// TIA Portal project "EMS" (V15.1) (continued)
   "SDC_EMS01_CARRIER61_Spare2" AT %Q6828.2 : Bool;
   "SDC_EMS01_CARRIER61_PositioningComplete" AT %Q6828.3 : Bool;
   "SDC_EMS01_CARRIER61_RunStopPressed" AT %Q6828.4 : Bool;
   "SDC_EMS01_CARRIER61_Moving" AT %Q6828.5 : Bool;
   "SDC_EMS01_CARRIER61_Faulted" AT %Q6828.6 : Bool;
   "SDC_EMS01_CARRIER61_InAuto" AT %Q6828.7 : Bool;
   "SDC_EMS01_CARRIER62_Spare0" AT %Q6829.0 : Bool;
   "SDC_EMS01_CARRIER62_DriveTripped" AT %Q6829.1 : Bool;
   "SDC_EMS01_CARRIER62_Spare2" AT %Q6829.2 : Bool;
   "SDC_EMS01_CARRIER62_PositioningComplete" AT %Q6829.3 : Bool;
   "SDC_EMS01_CARRIER62_RunStopPressed" AT %Q6829.4 : Bool;
   "SDC_EMS01_CARRIER62_Moving" AT %Q6829.5 : Bool;
   "SDC_EMS01_CARRIER62_Faulted" AT %Q6829.6 : Bool;
   "SDC_EMS01_CARRIER62_InAuto" AT %Q6829.7 : Bool;
   "SDC_EMS01_CARRIER63_Spare0" AT %Q6830.0 : Bool;
   "SDC_EMS01_CARRIER63_DriveTripped" AT %Q6830.1 : Bool;
   "SDC_EMS01_CARRIER63_Spare2" AT %Q6830.2 : Bool;
   "SDC_EMS01_CARRIER63_PositioningComplete" AT %Q6830.3 : Bool;
   "SDC_EMS01_CARRIER63_RunStopPressed" AT %Q6830.4 : Bool;
   "SDC_EMS01_CARRIER63_Moving" AT %Q6830.5 : Bool;
   "SDC_EMS01_CARRIER63_Faulted" AT %Q6830.6 : Bool;
   "SDC_EMS01_CARRIER63_InAuto" AT %Q6830.7 : Bool;
   "SDC_EMS01_CARRIER64_Spare0" AT %Q6831.0 : Bool;
   "SDC_EMS01_CARRIER64_DriveTripped" AT %Q6831.1 : Bool;
   "SDC_EMS01_CARRIER64_Spare2" AT %Q6831.2 : Bool;
   "SDC_EMS01_CARRIER64_PositioningComplete" AT %Q6831.3 : Bool;
   "SDC_EMS01_CARRIER64_RunStopPressed" AT %Q6831.4 : Bool;
   "SDC_EMS01_CARRIER64_Moving" AT %Q6831.5 : Bool;
   "SDC_EMS01_CARRIER64_Faulted" AT %Q6831.6 : Bool;
   "SDC_EMS01_CARRIER64_InAuto" AT %Q6831.7 : Bool;
   "SDC_EMS01_CARRIER65_Spare0" AT %Q6832.0 : Bool;
   "SDC_EMS01_CARRIER65_DriveTripped" AT %Q6832.1 : Bool;
   "SDC_EMS01_CARRIER65_Spare2" AT %Q6832.2 : Bool;
   "SDC_EMS01_CARRIER65_PositioningComplete" AT %Q6832.3 : Bool;
   "SDC_EMS01_CARRIER65_RunStopPressed" AT %Q6832.4 : Bool;
   "SDC_EMS01_CARRIER65_Moving" AT %Q6832.5 : Bool;
   "SDC_EMS01_CARRIER65_Faulted" AT %Q6832.6 : Bool;
   "SDC_EMS01_CARRIER65_InAuto" AT %Q6832.7 : Bool;
   "SDC_EMS01_CARRIER66_Spare0" AT %Q6833.0 : Bool;
   "SDC_EMS01_CARRIER66_DriveTripped" AT %Q6833.1 : Bool;
   "SDC_EMS01_CARRIER66_Spare2" AT %Q6833.2 : Bool;
   "SDC_EMS01_CARRIER66_PositioningComplete" AT %Q6833.3 : Bool;
   "SDC_EMS01_CARRIER66_RunStopPressed" AT %Q6833.4 : Bool;
   "SDC_EMS01_CARRIER66_Moving" AT %Q6833.5 : Bool;
   "SDC_EMS01_CARRIER66_Faulted" AT %Q6833.6 : Bool;
   "SDC_EMS01_CARRIER66_InAuto" AT %Q6833.7 : Bool;
   "SDC_EMS01_CARRIER67_Spare0" AT %Q6834.0 : Bool;
   "SDC_EMS01_CARRIER67_DriveTripped" AT %Q6834.1 : Bool;
   "SDC_EMS01_CARRIER67_Spare2" AT %Q6834.2 : Bool;
   "SDC_EMS01_CARRIER67_PositioningComplete" AT %Q6834.3 : Bool;
   "SDC_EMS01_CARRIER67_RunStopPressed" AT %Q6834.4 : Bool;
   "SDC_EMS01_CARRIER67_Moving" AT %Q6834.5 : Bool;
   "SDC_EMS01_CARRIER67_Faulted" AT %Q6834.6 : Bool;
   "SDC_EMS01_CARRIER67_InAuto" AT %Q6834.7 : Bool;
   "SDC_EMS01_CARRIER68_Spare0" AT %Q6835.0 : Bool;
   "SDC_EMS01_CARRIER68_DriveTripped" AT %Q6835.1 : Bool;
   "SDC_EMS01_CARRIER68_Spare2" AT %Q6835.2 : Bool;
   "SDC_EMS01_CARRIER68_PositioningComplete" AT %Q6835.3 : Bool;
   "SDC_EMS01_CARRIER68_RunStopPressed" AT %Q6835.4 : Bool;
   "SDC_EMS01_CARRIER68_Moving" AT %Q6835.5 : Bool;
   "SDC_EMS01_CARRIER68_Faulted" AT %Q6835.6 : Bool;
   "SDC_EMS01_CARRIER68_InAuto" AT %Q6835.7 : Bool;
   "SDC_EMS01_CARRIER69_Spare0" AT %Q6836.0 : Bool;
   "SDC_EMS01_CARRIER69_DriveTripped" AT %Q6836.1 : Bool;
   "SDC_EMS01_CARRIER69_Spare2" AT %Q6836.2 : Bool;
   "SDC_EMS01_CARRIER69_PositioningComplete" AT %Q6836.3 : Bool;
   "SDC_EMS01_CARRIER69_RunStopPressed" AT %Q6836.4 : Bool;
   "SDC_EMS01_CARRIER69_Moving" AT %Q6836.5 : Bool;
   "SDC_EMS01_CARRIER69_Faulted" AT %Q6836.6 : Bool;
   "SDC_EMS01_CARRIER69_InAuto" AT %Q6836.7 : Bool;
   "SDC_EMS01_CARRIER70_Spare0" AT %Q6837.0 : Bool;
   "SDC_EMS01_CARRIER70_DriveTripped" AT %Q6837.1 : Bool;
   "SDC_EMS01_CARRIER70_Spare2" AT %Q6837.2 : Bool;
   "SDC_EMS01_CARRIER70_PositioningComplete" AT %Q6837.3 : Bool;
   "SDC_EMS01_CARRIER70_RunStopPressed" AT %Q6837.4 : Bool;
   "SDC_EMS01_CARRIER70_Moving" AT %Q6837.5 : Bool;
   "SDC_EMS01_CARRIER70_Faulted" AT %Q6837.6 : Bool;
   "SDC_EMS01_CARRIER70_InAuto" AT %Q6837.7 : Bool;
   "SDC_EMS01_CARRIER71_Spare0" AT %Q6838.0 : Bool;
   "SDC_EMS01_CARRIER71_DriveTripped" AT %Q6838.1 : Bool;
   "SDC_EMS01_CARRIER71_Spare2" AT %Q6838.2 : Bool;
   "SDC_EMS01_CARRIER71_PositioningComplete" AT %Q6838.3 : Bool;
   "SDC_EMS01_CARRIER71_RunStopPressed" AT %Q6838.4 : Bool;
   "SDC_EMS01_CARRIER71_Moving" AT %Q6838.5 : Bool;
   "SDC_EMS01_CARRIER71_Faulted" AT %Q6838.6 : Bool;
   "SDC_EMS01_CARRIER71_InAuto" AT %Q6838.7 : Bool;
   "SDC_EMS01_CARRIER72_Spare0" AT %Q6839.0 : Bool;
   "SDC_EMS01_CARRIER72_DriveTripped" AT %Q6839.1 : Bool;
   "SDC_EMS01_CARRIER72_Spare2" AT %Q6839.2 : Bool;
   "SDC_EMS01_CARRIER72_PositioningComplete" AT %Q6839.3 : Bool;
   "SDC_EMS01_CARRIER72_RunStopPressed" AT %Q6839.4 : Bool;
   "SDC_EMS01_CARRIER72_Moving" AT %Q6839.5 : Bool;
   "SDC_EMS01_CARRIER72_Faulted" AT %Q6839.6 : Bool;
   "SDC_EMS01_CARRIER72_InAuto" AT %Q6839.7 : Bool;
   "SDC_EMS01_CARRIER73_Spare0" AT %Q6840.0 : Bool;
   "SDC_EMS01_CARRIER73_DriveTripped" AT %Q6840.1 : Bool;
   "SDC_EMS01_CARRIER73_Spare2" AT %Q6840.2 : Bool;
   "SDC_EMS01_CARRIER73_PositioningComplete" AT %Q6840.3 : Bool;
   "SDC_EMS01_CARRIER73_RunStopPressed" AT %Q6840.4 : Bool;
   "SDC_EMS01_CARRIER73_Moving" AT %Q6840.5 : Bool;
   "SDC_EMS01_CARRIER73_Faulted" AT %Q6840.6 : Bool;
   "SDC_EMS01_CARRIER73_InAuto" AT %Q6840.7 : Bool;
   "SDC_EMS01_CARRIER74_Spare0" AT %Q6841.0 : Bool;
   "SDC_EMS01_CARRIER74_DriveTripped" AT %Q6841.1 : Bool;
   "SDC_EMS01_CARRIER74_Spare2" AT %Q6841.2 : Bool;
   "SDC_EMS01_CARRIER74_PositioningComplete" AT %Q6841.3 : Bool;
   "SDC_EMS01_CARRIER74_RunStopPressed" AT %Q6841.4 : Bool;
   "SDC_EMS01_CARRIER74_Moving" AT %Q6841.5 : Bool;
   "SDC_EMS01_CARRIER74_Faulted" AT %Q6841.6 : Bool;
   "SDC_EMS01_CARRIER74_InAuto" AT %Q6841.7 : Bool;
   "SDC_EMS01_CARRIER75_Spare0" AT %Q6842.0 : Bool;
   "SDC_EMS01_CARRIER75_DriveTripped" AT %Q6842.1 : Bool;
   "SDC_EMS01_CARRIER75_Spare2" AT %Q6842.2 : Bool;
   "SDC_EMS01_CARRIER75_PositioningComplete" AT %Q6842.3 : Bool;
   "SDC_EMS01_CARRIER75_RunStopPressed" AT %Q6842.4 : Bool;
   "SDC_EMS01_CARRIER75_Moving" AT %Q6842.5 : Bool;
   "SDC_EMS01_CARRIER75_Faulted" AT %Q6842.6 : Bool;
   "SDC_EMS01_CARRIER75_InAuto" AT %Q6842.7 : Bool;
   "SDC_EMS01_CARRIER76_Spare0" AT %Q6843.0 : Bool;
   "SDC_EMS01_CARRIER76_DriveTripped" AT %Q6843.1 : Bool;
   "SDC_EMS01_CARRIER76_Spare2" AT %Q6843.2 : Bool;
   "SDC_EMS01_CARRIER76_PositioningComplete" AT %Q6843.3 : Bool;
   "SDC_EMS01_CARRIER76_RunStopPressed" AT %Q6843.4 : Bool;
   "SDC_EMS01_CARRIER76_Moving" AT %Q6843.5 : Bool;
   "SDC_EMS01_CARRIER76_Faulted" AT %Q6843.6 : Bool;
   "SDC_EMS01_CARRIER76_InAuto" AT %Q6843.7 : Bool;
   "SDC_EMS01_CARRIER77_Spare0" AT %Q6844.0 : Bool;
   "SDC_EMS01_CARRIER77_DriveTripped" AT %Q6844.1 : Bool;
   "SDC_EMS01_CARRIER77_Spare2" AT %Q6844.2 : Bool;
   "SDC_EMS01_CARRIER77_PositioningComplete" AT %Q6844.3 : Bool;
   "SDC_EMS01_CARRIER77_RunStopPressed" AT %Q6844.4 : Bool;
   "SDC_EMS01_CARRIER77_Moving" AT %Q6844.5 : Bool;
   "SDC_EMS01_CARRIER77_Faulted" AT %Q6844.6 : Bool;
   "SDC_EMS01_CARRIER77_InAuto" AT %Q6844.7 : Bool;
   "SDC_EMS01_CARRIER78_Spare0" AT %Q6845.0 : Bool;
   "SDC_EMS01_CARRIER78_DriveTripped" AT %Q6845.1 : Bool;
   "SDC_EMS01_CARRIER78_Spare2" AT %Q6845.2 : Bool;
   "SDC_EMS01_CARRIER78_PositioningComplete" AT %Q6845.3 : Bool;
   "SDC_EMS01_CARRIER78_RunStopPressed" AT %Q6845.4 : Bool;
   "SDC_EMS01_CARRIER78_Moving" AT %Q6845.5 : Bool;
   "SDC_EMS01_CARRIER78_Faulted" AT %Q6845.6 : Bool;
   "SDC_EMS01_CARRIER78_InAuto" AT %Q6845.7 : Bool;
   "SDC_EMS01_CARRIER79_Spare0" AT %Q6846.0 : Bool;
   "SDC_EMS01_CARRIER79_DriveTripped" AT %Q6846.1 : Bool;
   "SDC_EMS01_CARRIER79_Spare2" AT %Q6846.2 : Bool;
   "SDC_EMS01_CARRIER79_PositioningComplete" AT %Q6846.3 : Bool;
   "SDC_EMS01_CARRIER79_RunStopPressed" AT %Q6846.4 : Bool;
   "SDC_EMS01_CARRIER79_Moving" AT %Q6846.5 : Bool;
   "SDC_EMS01_CARRIER79_Faulted" AT %Q6846.6 : Bool;
   "SDC_EMS01_CARRIER79_InAuto" AT %Q6846.7 : Bool;
   "SDC_EMS01_CARRIER80_Spare0" AT %Q6847.0 : Bool;
   "SDC_EMS01_CARRIER80_DriveTripped" AT %Q6847.1 : Bool;
   "SDC_EMS01_CARRIER80_Spare2" AT %Q6847.2 : Bool;
   "SDC_EMS01_CARRIER80_PositioningComplete" AT %Q6847.3 : Bool;
   "SDC_EMS01_CARRIER80_RunStopPressed" AT %Q6847.4 : Bool;
   "SDC_EMS01_CARRIER80_Moving" AT %Q6847.5 : Bool;
   "SDC_EMS01_CARRIER80_Faulted" AT %Q6847.6 : Bool;
   "SDC_EMS01_CARRIER80_InAuto" AT %Q6847.7 : Bool;
   "SDC_EMS01_CARRIER81_Spare0" AT %Q6848.0 : Bool;
   "SDC_EMS01_CARRIER81_DriveTripped" AT %Q6848.1 : Bool;
   "SDC_EMS01_CARRIER81_Spare2" AT %Q6848.2 : Bool;
   "SDC_EMS01_CARRIER81_PositioningComplete" AT %Q6848.3 : Bool;
   "SDC_EMS01_CARRIER81_RunStopPressed" AT %Q6848.4 : Bool;
   "SDC_EMS01_CARRIER81_Moving" AT %Q6848.5 : Bool;
   "SDC_EMS01_CARRIER81_Faulted" AT %Q6848.6 : Bool;
   "SDC_EMS01_CARRIER81_InAuto" AT %Q6848.7 : Bool;
   "SDC_EMS01_CARRIER82_Spare0" AT %Q6849.0 : Bool;
   "SDC_EMS01_CARRIER82_DriveTripped" AT %Q6849.1 : Bool;
   "SDC_EMS01_CARRIER82_Spare2" AT %Q6849.2 : Bool;
   "SDC_EMS01_CARRIER82_PositioningComplete" AT %Q6849.3 : Bool;
   "SDC_EMS01_CARRIER82_RunStopPressed" AT %Q6849.4 : Bool;
   "SDC_EMS01_CARRIER82_Moving" AT %Q6849.5 : Bool;
   "SDC_EMS01_CARRIER82_Faulted" AT %Q6849.6 : Bool;
   "SDC_EMS01_CARRIER82_InAuto" AT %Q6849.7 : Bool;
   "SDC_EMS01_CARRIER83_Spare0" AT %Q6850.0 : Bool;
   "SDC_EMS01_CARRIER83_DriveTripped" AT %Q6850.1 : Bool;
   "SDC_EMS01_CARRIER83_Spare2" AT %Q6850.2 : Bool;
   "SDC_EMS01_CARRIER83_PositioningComplete" AT %Q6850.3 : Bool;
   "SDC_EMS01_CARRIER83_RunStopPressed" AT %Q6850.4 : Bool;
   "SDC_EMS01_CARRIER83_Moving" AT %Q6850.5 : Bool;
   "SDC_EMS01_CARRIER83_Faulted" AT %Q6850.6 : Bool;
   "SDC_EMS01_CARRIER83_InAuto" AT %Q6850.7 : Bool;
   "SDC_EMS01_CARRIER84_Spare0" AT %Q6851.0 : Bool;
   "SDC_EMS01_CARRIER84_DriveTripped" AT %Q6851.1 : Bool;
   "SDC_EMS01_CARRIER84_Spare2" AT %Q6851.2 : Bool;
   "SDC_EMS01_CARRIER84_PositioningComplete" AT %Q6851.3 : Bool;
   "SDC_EMS01_CARRIER84_RunStopPressed" AT %Q6851.4 : Bool;
   "SDC_EMS01_CARRIER84_Moving" AT %Q6851.5 : Bool;
   "SDC_EMS01_CARRIER84_Faulted" AT %Q6851.6 : Bool;
   "SDC_EMS01_CARRIER84_InAuto" AT %Q6851.7 : Bool;
   "SDC_EMS01_CARRIER85_Spare0" AT %Q6852.0 : Bool;
   "SDC_EMS01_CARRIER85_DriveTripped" AT %Q6852.1 : Bool;
   "SDC_EMS01_CARRIER85_Spare2" AT %Q6852.2 : Bool;
   "SDC_EMS01_CARRIER85_PositioningComplete" AT %Q6852.3 : Bool;
   "SDC_EMS01_CARRIER85_RunStopPressed" AT %Q6852.4 : Bool;
   "SDC_EMS01_CARRIER85_Moving" AT %Q6852.5 : Bool;
   "SDC_EMS01_CARRIER85_Faulted" AT %Q6852.6 : Bool;
   "SDC_EMS01_CARRIER85_InAuto" AT %Q6852.7 : Bool;
   "SDC_EMS01_CARRIER86_Spare0" AT %Q6853.0 : Bool;
   "SDC_EMS01_CARRIER86_DriveTripped" AT %Q6853.1 : Bool;
   "SDC_EMS01_CARRIER86_Spare2" AT %Q6853.2 : Bool;
   "SDC_EMS01_CARRIER86_PositioningComplete" AT %Q6853.3 : Bool;
   "SDC_EMS01_CARRIER86_RunStopPressed" AT %Q6853.4 : Bool;
   "SDC_EMS01_CARRIER86_Moving" AT %Q6853.5 : Bool;
   "SDC_EMS01_CARRIER86_Faulted" AT %Q6853.6 : Bool;
   "SDC_EMS01_CARRIER86_InAuto" AT %Q6853.7 : Bool;
   "SDC_EMS01_CARRIER87_Spare0" AT %Q6854.0 : Bool;
   "SDC_EMS01_CARRIER87_DriveTripped" AT %Q6854.1 : Bool;
   "SDC_EMS01_CARRIER87_Spare2" AT %Q6854.2 : Bool;
   "SDC_EMS01_CARRIER87_PositioningComplete" AT %Q6854.3 : Bool;
   "SDC_EMS01_CARRIER87_RunStopPressed" AT %Q6854.4 : Bool;
   "SDC_EMS01_CARRIER87_Moving" AT %Q6854.5 : Bool;
   "SDC_EMS01_CARRIER87_Faulted" AT %Q6854.6 : Bool;
   "SDC_EMS01_CARRIER87_InAuto" AT %Q6854.7 : Bool;
   "SDC_EMS01_CARRIER88_Spare0" AT %Q6855.0 : Bool;
   "SDC_EMS01_CARRIER88_DriveTripped" AT %Q6855.1 : Bool;
   "SDC_EMS01_CARRIER88_Spare2" AT %Q6855.2 : Bool;
   "SDC_EMS01_CARRIER88_PositioningComplete" AT %Q6855.3 : Bool;
   "SDC_EMS01_CARRIER88_RunStopPressed" AT %Q6855.4 : Bool;
   "SDC_EMS01_CARRIER88_Moving" AT %Q6855.5 : Bool;
   "SDC_EMS01_CARRIER88_Faulted" AT %Q6855.6 : Bool;
   "SDC_EMS01_CARRIER88_InAuto" AT %Q6855.7 : Bool;
   "SDC_EMS01_CARRIER89_Spare0" AT %Q6856.0 : Bool;
   "SDC_EMS01_CARRIER89_DriveTripped" AT %Q6856.1 : Bool;
   "SDC_EMS01_CARRIER89_Spare2" AT %Q6856.2 : Bool;
   "SDC_EMS01_CARRIER89_PositioningComplete" AT %Q6856.3 : Bool;
   "SDC_EMS01_CARRIER89_RunStopPressed" AT %Q6856.4 : Bool;
   "SDC_EMS01_CARRIER89_Moving" AT %Q6856.5 : Bool;
   "SDC_EMS01_CARRIER89_Faulted" AT %Q6856.6 : Bool;
   "SDC_EMS01_CARRIER89_InAuto" AT %Q6856.7 : Bool;
   "SDC_EMS01_CARRIER90_Spare0" AT %Q6857.0 : Bool;
   "SDC_EMS01_CARRIER90_DriveTripped" AT %Q6857.1 : Bool;
   "SDC_EMS01_CARRIER90_Spare2" AT %Q6857.2 : Bool;
   "SDC_EMS01_CARRIER90_PositioningComplete" AT %Q6857.3 : Bool;
   "SDC_EMS01_CARRIER90_RunStopPressed" AT %Q6857.4 : Bool;
   "SDC_EMS01_CARRIER90_Moving" AT %Q6857.5 : Bool;
   "SDC_EMS01_CARRIER90_Faulted" AT %Q6857.6 : Bool;
   "SDC_EMS01_CARRIER90_InAuto" AT %Q6857.7 : Bool;
   "SDC_EMS01_CARRIER91_Spare0" AT %Q6858.0 : Bool;
   "SDC_EMS01_CARRIER91_DriveTripped" AT %Q6858.1 : Bool;
   "SDC_EMS01_CARRIER91_Spare2" AT %Q6858.2 : Bool;
   "SDC_EMS01_CARRIER91_PositioningComplete" AT %Q6858.3 : Bool;
   "SDC_EMS01_CARRIER91_RunStopPressed" AT %Q6858.4 : Bool;
   "SDC_EMS01_CARRIER91_Moving" AT %Q6858.5 : Bool;
   "SDC_EMS01_CARRIER91_Faulted" AT %Q6858.6 : Bool;
   "SDC_EMS01_CARRIER91_InAuto" AT %Q6858.7 : Bool;
   "SDC_EMS01_CARRIER92_Spare0" AT %Q6859.0 : Bool;
   "SDC_EMS01_CARRIER92_DriveTripped" AT %Q6859.1 : Bool;
   "SDC_EMS01_CARRIER92_Spare2" AT %Q6859.2 : Bool;
   "SDC_EMS01_CARRIER92_PositioningComplete" AT %Q6859.3 : Bool;
   "SDC_EMS01_CARRIER92_RunStopPressed" AT %Q6859.4 : Bool;
   "SDC_EMS01_CARRIER92_Moving" AT %Q6859.5 : Bool;
   "SDC_EMS01_CARRIER92_Faulted" AT %Q6859.6 : Bool;
   "SDC_EMS01_CARRIER92_InAuto" AT %Q6859.7 : Bool;
   "SDC_EMS01_CARRIER93_Spare0" AT %Q6860.0 : Bool;
   "SDC_EMS01_CARRIER93_DriveTripped" AT %Q6860.1 : Bool;
   "SDC_EMS01_CARRIER93_Spare2" AT %Q6860.2 : Bool;
   "SDC_EMS01_CARRIER93_PositioningComplete" AT %Q6860.3 : Bool;
   "SDC_EMS01_CARRIER93_RunStopPressed" AT %Q6860.4 : Bool;
   "SDC_EMS01_CARRIER93_Moving" AT %Q6860.5 : Bool;
   "SDC_EMS01_CARRIER93_Faulted" AT %Q6860.6 : Bool;
   "SDC_EMS01_CARRIER93_InAuto" AT %Q6860.7 : Bool;
   "SDC_EMS01_CARRIER94_Spare0" AT %Q6861.0 : Bool;
   "SDC_EMS01_CARRIER94_DriveTripped" AT %Q6861.1 : Bool;
   "SDC_EMS01_CARRIER94_Spare2" AT %Q6861.2 : Bool;
   "SDC_EMS01_CARRIER94_PositioningComplete" AT %Q6861.3 : Bool;
   "SDC_EMS01_CARRIER94_RunStopPressed" AT %Q6861.4 : Bool;
   "SDC_EMS01_CARRIER94_Moving" AT %Q6861.5 : Bool;
   "SDC_EMS01_CARRIER94_Faulted" AT %Q6861.6 : Bool;
   "SDC_EMS01_CARRIER94_InAuto" AT %Q6861.7 : Bool;
   "SDC_EMS01_CARRIER95_Spare0" AT %Q6862.0 : Bool;
   "SDC_EMS01_CARRIER95_DriveTripped" AT %Q6862.1 : Bool;
   "SDC_EMS01_CARRIER95_Spare2" AT %Q6862.2 : Bool;
   "SDC_EMS01_CARRIER95_PositioningComplete" AT %Q6862.3 : Bool;
   "SDC_EMS01_CARRIER95_RunStopPressed" AT %Q6862.4 : Bool;
   "SDC_EMS01_CARRIER95_Moving" AT %Q6862.5 : Bool;
   "SDC_EMS01_CARRIER95_Faulted" AT %Q6862.6 : Bool;
   "SDC_EMS01_CARRIER95_InAuto" AT %Q6862.7 : Bool;
   "EMS01_MASTER_POWER_ON_ON_DELAY_" AT %I6000.0 : Bool;
   "EMS01_FAULT_RESET__PB_2406" AT %I6000.1 : Bool;
   "EMS01R1_MASTER_POWER_ON_ON_DELAY_" AT %I6000.2 : Bool;
   "EMS01R1_FAULT_RESET__PB_2406" AT %I6000.3 : Bool;
   "EMS01R2_MASTER_POWER_ON_ON_DELAY_" AT %I6000.4 : Bool;
   "EMS01R2_FAULT_RESET__PB_2406" AT %I6000.5 : Bool;
   "EMS01R3_MASTER_POWER_ON_ON_DELAY_" AT %I6000.6 : Bool;
   "EMS01R3_FAULT_RESET__PB_2406" AT %I6000.7 : Bool;
   "EMS01R4_MASTER_POWER_ON_ON_DELAY_" AT %I6001.0 : Bool;
   "EMS01R4_FAULT_RESET__PB_3206" AT %I6001.1 : Bool;
   "Stop_#26__Set_To_Release" AT %I6001.2 : Bool;
   "SPARE_EMS_TO_SDC" AT %I6001.3 : Bool;
   "SPARE_EMS_TO_SDC(1)" AT %I6001.4 : Bool;
   "SPARE_EMS_TO_SDC(2)" AT %I6001.5 : Bool;
   "SPARE_EMS_TO_SDC(3)" AT %I6001.6 : Bool;
   "Heartbeat" AT %I6001.7 : Bool;
   "SPARE_EMS_TO_SDC(4)" AT %IW6002 : Word;
   "SPARE_EMS_TO_SDC(5)" AT %IW6004 : Word;
   "CARRIER_SPEED" AT %IW6006 : Word;
   "PRODUCTION_SPEED_REF_MM_MIN" AT %IW6008 : Word;
   "PRODUCTION_SPEED_REF_FT_MIN" AT %IW6010 : Word;
   "Speed_Thru_Test_Zone" AT %IW6012 : Word;
   "PANELVIEW_#1_CARRIER_SELECTED_TO_BE_DELETED" AT %IW6014 : Word;
   "PANELVIEW_#2_CARRIER_SELECTED_TO_BE_DELETED" AT %IW6016 : Word;
   "PANELVIEW_#3_CARRIER_SELECTED_TO_BE_DELETED" AT %IW6018 : Word;
   "PANELVIEW_#4_CARRIER_SELECTED_TO_BE_DELETED" AT %IW6020 : Word;
   "PANELVIEW_#5_CARRIER_SELECTED_TO_BE_DELETED" AT %IW6022 : Word;
   "PANELVIEW_#6_CARRIER_SELECTED_TO_BE_DELETED" AT %IW6024 : Word;
   "SPARE_EMS_TO_SDC(6)" AT %IW6026 : Word;
   "SPARE_EMS_TO_SDC(7)" AT %IW6028 : Word;
   "STOP1_CONTROL_FROM_EMS01" AT %ID6030 : DWord;
   "STOP2_CONTROL_FROM_EMS01" AT %ID6034 : DWord;
   "STOP3_CONTROL_FROM_EMS01" AT %ID6038 : DWord;
   "STOP4_CONTROL_FROM_EMS01" AT %ID6042 : DWord;
   "STOP5_CONTROL_FROM_EMS01" AT %ID6046 : DWord;
   "STOP6_CONTROL_FROM_EMS01" AT %ID6050 : DWord;
   "STOP7_CONTROL_FROM_EMS01" AT %ID6054 : DWord;
   "STOP8_CONTROL_FROM_EMS01" AT %ID6058 : DWord;
   "STOP9_CONTROL_FROM_EMS01" AT %ID6062 : DWord;
   "STOP10_CONTROL_FROM_EMS01" AT %ID6066 : DWord;
   "STOP11_CONTROL_FROM_EMS01" AT %ID6070 : DWord;
   "STOP12_CONTROL_FROM_EMS01" AT %ID6074 : DWord;
   "STOP13_CONTROL_FROM_EMS01" AT %ID6078 : DWord;
   "STOP14_CONTROL_FROM_EMS01" AT %ID6082 : DWord;
   "STOP15_CONTROL_FROM_EMS01" AT %ID6086 : DWord;
   "STOP16_CONTROL_FROM_EMS01" AT %ID6090 : DWord;
   "STOP17_CONTROL_FROM_EMS01" AT %ID6094 : DWord;
   "STOP18_CONTROL_FROM_EMS01" AT %ID6098 : DWord;
   "STOP19_CONTROL_FROM_EMS01" AT %ID6102 : DWord;
   "STOP20_CONTROL_FROM_EMS01" AT %ID6106 : DWord;
   "STOP21_CONTROL_FROM_EMS01" AT %ID6110 : DWord;
   "STOP22_CONTROL_FROM_EMS01" AT %ID6114 : DWord;
   "STOP23_CONTROL_FROM_EMS01" AT %ID6118 : DWord;
   "STOP24_CONTROL_FROM_EMS01" AT %ID6122 : DWord;
   "STOP25_CONTROL_FROM_EMS01" AT %ID6126 : DWord;
   "STOP26_CONTROL_FROM_EMS01" AT %ID6130 : DWord;
   "STOP27_CONTROL_FROM_EMS01" AT %ID6134 : DWord;
   "STOP28_CONTROL_FROM_EMS01" AT %ID6138 : DWord;
   "STOP29_CONTROL_FROM_EMS01" AT %ID6142 : DWord;
   "STOP30_CONTROL_FROM_EMS01" AT %ID6146 : DWord;
   "STOP31_CONTROL_FROM_EMS01" AT %ID6150 : DWord;
   "STOP32_CONTROL_FROM_EMS01" AT %ID6154 : DWord;
   "STOP33_CONTROL_FROM_EMS01" AT %ID6158 : DWord;
   "STOP34_CONTROL_FROM_EMS01" AT %ID6162 : DWord;
   "STOP35_CONTROL_FROM_EMS01" AT %ID6166 : DWord;
   "STOP36_CONTROL_FROM_EMS01" AT %ID6170 : DWord;
   "STOP37_CONTROL_FROM_EMS01" AT %ID6174 : DWord;
   "STOP38_CONTROL_FROM_EMS01" AT %ID6178 : DWord;
   "STOP39_CONTROL_FROM_EMS01" AT %ID6182 : DWord;
   "STOP40_CONTROL_FROM_EMS01" AT %ID6186 : DWord;
   "STOP41_CONTROL_FROM_EMS01" AT %ID6190 : DWord;
   "STOP42_CONTROL_FROM_EMS01" AT %ID6194 : DWord;
   "STOP43_CONTROL_FROM_EMS01" AT %ID6198 : DWord;
   "STOP44_CONTROL_FROM_EMS01" AT %ID6202 : DWord;
   "STOP45_CONTROL_FROM_EMS01" AT %ID6206 : DWord;
   "STOP46_CONTROL_FROM_EMS01" AT %ID6210 : DWord;
   "STOP47_CONTROL_FROM_EMS01" AT %ID6214 : DWord;
   "STOP48_CONTROL_FROM_EMS01" AT %ID6218 : DWord;
   "STOP49_CONTROL_FROM_EMS01" AT %ID6222 : DWord;
   "STOP50_CONTROL_FROM_EMS01" AT %ID6226 : DWord;
   "STOP51_CONTROL_FROM_EMS01" AT %ID6230 : DWord;
   "STOP52_CONTROL_FROM_EMS01" AT %ID6234 : DWord;
   "STOP53_CONTROL_FROM_EMS01" AT %ID6238 : DWord;
   "STOP54_CONTROL_FROM_EMS01" AT %ID6242 : DWord;
   "STOP55_CONTROL_FROM_EMS01" AT %ID6246 : DWord;
   "STOP56_CONTROL_FROM_EMS01" AT %ID6250 : DWord;
   "STOP57_CONTROL_FROM_EMS01" AT %ID6254 : DWord;
   "STOP58_CONTROL_FROM_EMS01" AT %ID6258 : DWord;
   "STOP59_CONTROL_FROM_EMS01" AT %ID6262 : DWord;
   "STOP60_CONTROL_FROM_EMS01" AT %ID6266 : DWord;
   "STOP61_CONTROL_FROM_EMS01" AT %ID6270 : DWord;
   "STOP62_CONTROL_FROM_EMS01" AT %ID6274 : DWord;
   "STOP63_CONTROL_FROM_EMS01" AT %ID6278 : DWord;
   "STOP64_CONTROL_FROM_EMS01" AT %ID6282 : DWord;
   "STOP65_CONTROL_FROM_EMS01" AT %ID6286 : DWord;
   "SPARE" AT %ID6290 : DWord;
   "SPARE(1)" AT %ID6294 : DWord;
   "SPARE(2)" AT %ID6298 : DWord;
   "SPARE(3)" AT %ID6302 : DWord;
   "SPARE(4)" AT %ID6306 : DWord;
   "SPARE(5)" AT %ID6310 : DWord;
   "SPARE(6)" AT %ID6314 : DWord;
   "SPARE(7)" AT %ID6318 : DWord;
   "SPARE(8)" AT %ID6322 : DWord;
   "SPARE(9)" AT %ID6326 : DWord;
   "SPARE(10)" AT %ID6330 : DWord;
   "SPARE(11)" AT %ID6334 : DWord;
   "SPARE(12)" AT %ID6338 : DWord;
   "SPARE(13)" AT %ID6342 : DWord;
   "SPARE(14)" AT %ID6346 : DWord;
   "SDC_EMS01_Carrier1_Fault" AT %QB7024 : Byte;
   "SDC_EMS01_Carrier2_Fault" AT %QB7025 : Byte;
   "SDC_EMS01_Carrier3_Fault" AT %QB7026 : Byte;
   "SDC_EMS01_Carrier4_Fault" AT %QB7027 : Byte;
   "SDC_EMS01_Carrier5_Fault" AT %QB7028 : Byte;
   "SDC_EMS01_Carrier6_Fault" AT %QB7029 : Byte;
   "SDC_EMS01_Carrier7_Fault" AT %QB7030 : Byte;
   "SDC_EMS01_Carrier8_Fault" AT %QB7031 : Byte;
   "SDC_EMS01_Carrier9_Fault" AT %QB7032 : Byte;
   "SDC_EMS01_Carrier10_Fault" AT %QB7033 : Byte;
   "SDC_EMS01_Carrier11_Fault" AT %QB7034 : Byte;
   "SDC_EMS01_Carrier12_Fault" AT %QB7035 : Byte;
   "SDC_EMS01_Carrier13_Fault" AT %QB7036 : Byte;
   "SDC_EMS01_Carrier14_Fault" AT %QB7037 : Byte;
   "SDC_EMS01_Carrier15_Fault" AT %QB7038 : Byte;
   "SDC_EMS01_Carrier16_Fault" AT %QB7039 : Byte;
   "SDC_EMS01_Carrier17_Fault" AT %QB7040 : Byte;
   "SDC_EMS01_Carrier18_Fault" AT %QB7041 : Byte;
   "SDC_EMS01_Carrier19_Fault" AT %QB7042 : Byte;
   "SDC_EMS01_Carrier20_Fault" AT %QB7043 : Byte;
   "SDC_EMS01_Carrier21_Fault" AT %QB7044 : Byte;
   "SDC_EMS01_Carrier22_Fault" AT %QB7045 : Byte;
   "SDC_EMS01_Carrier23_Fault" AT %QB7046 : Byte;
   "SDC_EMS01_Carrier24_Fault" AT %QB7047 : Byte;
   "SDC_EMS01_Carrier25_Fault" AT %QB7048 : Byte;
   "SDC_EMS01_Carrier26_Fault" AT %QB7049 : Byte;
   "SDC_EMS01_Carrier27_Fault" AT %QB7050 : Byte;
   "SDC_EMS01_Carrier28_Fault" AT %QB7051 : Byte;
   "SDC_EMS01_Carrier29_Fault" AT %QB7052 : Byte;
   "SDC_EMS01_Carrier30_Fault" AT %QB7053 : Byte;
   "SDC_EMS01_Carrier31_Fault" AT %QB7054 : Byte;
   "SDC_EMS01_Carrier32_Fault" AT %QB7055 : Byte;
   "SDC_EMS01_Carrier33_Fault" AT %QB7056 : Byte;
   "SDC_EMS01_Carrier34_Fault" AT %QB7057 : Byte;
   "SDC_EMS01_Carrier35_Fault" AT %QB7058 : Byte;
   "SDC_EMS01_Carrier36_Fault" AT %QB7059 : Byte;
   "SDC_EMS01_Carrier37_Fault" AT %QB7060 : Byte;
   "SDC_EMS01_Carrier38_Fault" AT %QB7061 : Byte;
   "SDC_EMS01_Carrier39_Fault" AT %QB7062 : Byte;
   "SDC_EMS01_Carrier40_Fault" AT %QB7063 : Byte;
   "SDC_EMS01_Carrier41_Fault" AT %QB7064 : Byte;
   "SDC_EMS01_Carrier42_Fault" AT %QB7065 : Byte;
   "SDC_EMS01_Carrier43_Fault" AT %QB7066 : Byte;
   "SDC_EMS01_Carrier44_Fault" AT %QB7067 : Byte;
   "SDC_EMS01_Carrier45_Fault" AT %QB7068 : Byte;
   "SDC_EMS01_Carrier46_Fault" AT %QB7069 : Byte;
   "SDC_EMS01_Carrier47_Fault" AT %QB7070 : Byte;
   "SDC_EMS01_Carrier48_Fault" AT %QB7071 : Byte;
   "SDC_EMS01_Carrier49_Fault" AT %QB7072 : Byte;
   "SDC_EMS01_Carrier50_Fault" AT %QB7073 : Byte;
   "SDC_EMS01_Carrier51_Fault" AT %QB7074 : Byte;
   "SDC_EMS01_Carrier52_Fault" AT %QB7075 : Byte;
   "SDC_EMS01_Carrier53_Fault" AT %QB7076 : Byte;
   "SDC_EMS01_Carrier54_Fault" AT %QB7077 : Byte;
   "SDC_EMS01_Carrier55_Fault" AT %QB7078 : Byte;
   "SDC_EMS01_Carrier56_Fault" AT %QB7079 : Byte;
   "SDC_EMS01_Carrier57_Fault" AT %QB7080 : Byte;
   "SDC_EMS01_Carrier58_Fault" AT %QB7081 : Byte;
   "SDC_EMS01_Carrier59_Fault" AT %QB7082 : Byte;
   "SDC_EMS01_Carrier60_Fault" AT %QB7083 : Byte;
   "SDC_EMS01_Carrier61_Fault" AT %QB7084 : Byte;
   "SDC_EMS01_Carrier62_Fault" AT %QB7085 : Byte;
   "SDC_EMS01_Carrier63_Fault" AT %QB7086 : Byte;
   "SDC_EMS01_Carrier64_Fault" AT %QB7087 : Byte;
   "SDC_EMS01_Carrier65_Fault" AT %QB7088 : Byte;
   "SDC_EMS01_Carrier66_Fault" AT %QB7089 : Byte;
   "SDC_EMS01_Carrier67_Fault" AT %QB7090 : Byte;
   "SDC_EMS01_Carrier68_Fault" AT %QB7091 : Byte;
   "SDC_EMS01_Carrier69_Fault" AT %QB7092 : Byte;
   "SDC_EMS01_Carrier70_Fault" AT %QB7093 : Byte;
   "SDC_EMS01_Carrier71_Fault" AT %QB7094 : Byte;
   "SDC_EMS01_Carrier72_Fault" AT %QB7095 : Byte;
   "SDC_EMS01_Carrier73_Fault" AT %QB7096 : Byte;
   "SDC_EMS01_Carrier74_Fault" AT %QB7097 : Byte;
   "SDC_EMS01_Carrier75_Fault" AT %QB7098 : Byte;
   "SDC_EMS01_Carrier76_Fault" AT %QB7099 : Byte;
   "SDC_EMS01_Carrier77_Fault" AT %QB7100 : Byte;
   "SDC_EMS01_Carrier78_Fault" AT %QB7101 : Byte;
   "SDC_EMS01_Carrier79_Fault" AT %QB7102 : Byte;
   "SDC_EMS01_Carrier80_Fault" AT %QB7103 : Byte;
   "SDC_EMS01_Carrier81_Fault" AT %QB7104 : Byte;
   "SDC_EMS01_Carrier82_Fault" AT %QB7105 : Byte;
   "SDC_EMS01_Carrier83_Fault" AT %QB7106 : Byte;
   "SDC_EMS01_Carrier84_Fault" AT %QB7107 : Byte;
   "SDC_EMS01_Carrier85_Fault" AT %QB7108 : Byte;
   "SDC_EMS01_Carrier86_Fault" AT %QB7109 : Byte;
   "SDC_EMS01_Carrier87_Fault" AT %QB7110 : Byte;
   "SDC_EMS01_Carrier88_Fault" AT %QB7111 : Byte;
   "SDC_EMS01_Carrier89_Fault" AT %QB7112 : Byte;
   "SDC_EMS01_Carrier90_Fault" AT %QB7113 : Byte;
   "SDC_EMS01_Carrier91_Fault" AT %QB7114 : Byte;
   "SDC_EMS01_Carrier92_Fault" AT %QB7115 : Byte;
   "SDC_EMS01_Carrier93_Fault" AT %QB7116 : Byte;
   "SDC_EMS01_Carrier94_Fault" AT %QB7117 : Byte;
   "SDC_EMS01_Carrier95_Fault" AT %QB7118 : Byte;
   "SDC_EMS01_Carrier1_status" AT %QB6768 : Byte;
   "SDC_EMS01_Carrier2_status" AT %QB6769 : Byte;
   "SDC_EMS01_Carrier3_status" AT %QB6770 : Byte;
   "SDC_EMS01_Carrier4_status" AT %QB6771 : Byte;
   "SDC_EMS01_Carrier5_status" AT %QB6772 : Byte;
   "SDC_EMS01_Carrier6_status" AT %QB6773 : Byte;
   "SDC_EMS01_Carrier7_status" AT %QB6774 : Byte;
   "SDC_EMS01_Carrier8_status" AT %QB6775 : Byte;
   "SDC_EMS01_Carrier9_status" AT %QB6776 : Byte;
   "SDC_EMS01_Carrier10_status" AT %QB6777 : Byte;
   "SDC_EMS01_Carrier11_status" AT %QB6778 : Byte;
   "SDC_EMS01_Carrier12_status" AT %QB6779 : Byte;
   "SDC_EMS01_Carrier13_status" AT %QB6780 : Byte;
   "SDC_EMS01_Carrier14_status" AT %QB6781 : Byte;
   "SDC_EMS01_Carrier15_status" AT %QB6782 : Byte;
   "SDC_EMS01_Carrier16_status" AT %QB6783 : Byte;
   "SDC_EMS01_Carrier17_status" AT %QB6784 : Byte;
   "SDC_EMS01_Carrier18_status" AT %QB6785 : Byte;
   "SDC_EMS01_Carrier19_status" AT %QB6786 : Byte;
   "SDC_EMS01_Carrier20_status" AT %QB6787 : Byte;
   "SDC_EMS01_Carrier21_status" AT %QB6788 : Byte;
   "SDC_EMS01_Carrier22_status" AT %QB6789 : Byte;
   "SDC_EMS01_Carrier23_status" AT %QB6790 : Byte;
   "SDC_EMS01_Carrier24_status" AT %QB6791 : Byte;
   "SDC_EMS01_Carrier25_status" AT %QB6792 : Byte;
   "SDC_EMS01_Carrier26_status" AT %QB6793 : Byte;
   "SDC_EMS01_Carrier27_status" AT %QB6794 : Byte;
   "SDC_EMS01_Carrier28_status" AT %QB6795 : Byte;
   "SDC_EMS01_Carrier29_status" AT %QB6796 : Byte;
   "SDC_EMS01_Carrier30_status" AT %QB6797 : Byte;
   "SDC_EMS01_Carrier31_status" AT %QB6798 : Byte;
   "SDC_EMS01_Carrier32_status" AT %QB6799 : Byte;
   "SDC_EMS01_Carrier33_status" AT %QB6800 : Byte;
   "SDC_EMS01_Carrier34_status" AT %QB6801 : Byte;
   "SDC_EMS01_Carrier35_status" AT %QB6802 : Byte;
   "SDC_EMS01_Carrier36_status" AT %QB6803 : Byte;
   "SDC_EMS01_Carrier37_status" AT %QB6804 : Byte;
   "SDC_EMS01_Carrier38_status" AT %QB6805 : Byte;
   "SDC_EMS01_Carrier39_status" AT %QB6806 : Byte;
   "SDC_EMS01_Carrier40_status" AT %QB6807 : Byte;
   "SDC_EMS01_Carrier41_status" AT %QB6808 : Byte;
   "SDC_EMS01_Carrier42_status" AT %QB6809 : Byte;
   "SDC_EMS01_Carrier43_status" AT %QB6810 : Byte;
   "SDC_EMS01_Carrier44_status" AT %QB6811 : Byte;
   "SDC_EMS01_Carrier45_status" AT %QB6812 : Byte;
   "SDC_EMS01_Carrier46_status" AT %QB6813 : Byte;
   "SDC_EMS01_Carrier47_status" AT %QB6814 : Byte;
   "SDC_EMS01_Carrier48_status" AT %QB6815 : Byte;
   "SDC_EMS01_Carrier49_status" AT %QB6816 : Byte;
   "SDC_EMS01_Carrier50_status" AT %QB6817 : Byte;
   "SDC_EMS01_Carrier51_status" AT %QB6818 : Byte;
   "SDC_EMS01_Carrier52_status" AT %QB6819 : Byte;
   "SDC_EMS01_Carrier53_status" AT %QB6820 : Byte;
   "SDC_EMS01_Carrier54_status" AT %QB6821 : Byte;
   "SDC_EMS01_Carrier55_status" AT %QB6822 : Byte;
   "SDC_EMS01_Carrier56_status" AT %QB6823 : Byte;
   "SDC_EMS01_Carrier57_status" AT %QB6824 : Byte;
   "SDC_EMS01_Carrier58_status" AT %QB6825 : Byte;
   "SDC_EMS01_Carrier59_status" AT %QB6826 : Byte;
   "SDC_EMS01_Carrier60_status" AT %QB6827 : Byte;
   "SDC_EMS01_Carrier61_status" AT %QB6828 : Byte;
   "SDC_EMS01_Carrier62_status" AT %QB6829 : Byte;
   "SDC_EMS01_Carrier63_status" AT %QB6830 : Byte;
   "SDC_EMS01_Carrier64_status" AT %QB6831 : Byte;
   "SDC_EMS01_Carrier65_status" AT %QB6832 : Byte;
   "SDC_EMS01_Carrier66_status" AT %QB6833 : Byte;
   "SDC_EMS01_Carrier67_status" AT %QB6834 : Byte;
   "SDC_EMS01_Carrier68_status" AT %QB6835 : Byte;
   "SDC_EMS01_Carrier69_status" AT %QB6836 : Byte;
   "SDC_EMS01_Carrier70_status" AT %QB6837 : Byte;
   "SDC_EMS01_Carrier71_status" AT %QB6838 : Byte;
   "SDC_EMS01_Carrier72_status" AT %QB6839 : Byte;
   "SDC_EMS01_Carrier73_status" AT %QB6840 : Byte;
   "SDC_EMS01_Carrier74_status" AT %QB6841 : Byte;
   "SDC_EMS01_Carrier75_status" AT %QB6842 : Byte;
   "SDC_EMS01_Carrier76_status" AT %QB6843 : Byte;
   "SDC_EMS01_Carrier77_status" AT %QB6844 : Byte;
   "SDC_EMS01_Carrier78_status" AT %QB6845 : Byte;
   "SDC_EMS01_Carrier79_status" AT %QB6846 : Byte;
   "SDC_EMS01_Carrier80_status" AT %QB6847 : Byte;
   "SDC_EMS01_Carrier81_status" AT %QB6848 : Byte;
   "SDC_EMS01_Carrier82_status" AT %QB6849 : Byte;
   "SDC_EMS01_Carrier83_status" AT %QB6850 : Byte;
   "SDC_EMS01_Carrier84_status" AT %QB6851 : Byte;
   "SDC_EMS01_Carrier85_status" AT %QB6852 : Byte;
   "SDC_EMS01_Carrier86_status" AT %QB6853 : Byte;
   "SDC_EMS01_Carrier87_status" AT %QB6854 : Byte;
   "SDC_EMS01_Carrier88_status" AT %QB6855 : Byte;
   "SDC_EMS01_Carrier89_status" AT %QB6856 : Byte;
   "SDC_EMS01_Carrier90_status" AT %QB6857 : Byte;
   "SDC_EMS01_Carrier91_status" AT %QB6858 : Byte;
   "SDC_EMS01_Carrier92_status" AT %QB6859 : Byte;
   "SDC_EMS01_Carrier93_status" AT %QB6860 : Byte;
   "SDC_EMS01_Carrier94_status" AT %QB6861 : Byte;
   "SDC_EMS01_Carrier95_status" AT %QB6862 : Byte;
   "SDC_EMS01_Carrier1_Zone" AT %QB6512 : Byte;
   "SDC_EMS01_Carrier2_Zone" AT %QB6513 : Byte;
   "SDC_EMS01_Carrier3_Zone" AT %QB6514 : Byte;
   "SDC_EMS01_Carrier4_Zone" AT %QB6515 : Byte;
   "SDC_EMS01_Carrier5_Zone" AT %QB6516 : Byte;
   "SDC_EMS01_Carrier6_Zone" AT %QB6517 : Byte;
   "SDC_EMS01_Carrier7_Zone" AT %QB6518 : Byte;
   "SDC_EMS01_Carrier8_Zone" AT %QB6519 : Byte;
   "SDC_EMS01_Carrier9_Zone" AT %QB6520 : Byte;
   "SDC_EMS01_Carrier10_Zone" AT %QB6521 : Byte;
   "SDC_EMS01_Carrier11_Zone" AT %QB6522 : Byte;
   "SDC_EMS01_Carrier12_Zone" AT %QB6523 : Byte;
   "SDC_EMS01_Carrier13_Zone" AT %QB6524 : Byte;
   "SDC_EMS01_Carrier14_Zone" AT %QB6525 : Byte;
   "SDC_EMS01_Carrier15_Zone" AT %QB6526 : Byte;
   "SDC_EMS01_Carrier16_Zone" AT %QB6527 : Byte;
   "SDC_EMS01_Carrier17_Zone" AT %QB6528 : Byte;
   "SDC_EMS01_Carrier18_Zone" AT %QB6529 : Byte;
   "SDC_EMS01_Carrier19_Zone" AT %QB6530 : Byte;
   "SDC_EMS01_Carrier20_Zone" AT %QB6531 : Byte;
   "SDC_EMS01_Carrier21_Zone" AT %QB6532 : Byte;
   "SDC_EMS01_Carrier22_Zone" AT %QB6533 : Byte;
   "SDC_EMS01_Carrier23_Zone" AT %QB6534 : Byte;
   "SDC_EMS01_Carrier24_Zone" AT %QB6535 : Byte;
   "SDC_EMS01_Carrier25_Zone" AT %QB6536 : Byte;
   "SDC_EMS01_Carrier26_Zone" AT %QB6537 : Byte;
   "SDC_EMS01_Carrier27_Zone" AT %QB6538 : Byte;
   "SDC_EMS01_Carrier28_Zone" AT %QB6539 : Byte;
   "SDC_EMS01_Carrier29_Zone" AT %QB6540 : Byte;
   "SDC_EMS01_Carrier30_Zone" AT %QB6541 : Byte;
   "SDC_EMS01_Carrier31_Zone" AT %QB6542 : Byte;
   "SDC_EMS01_Carrier32_Zone" AT %QB6543 : Byte;
   "SDC_EMS01_Carrier33_Zone" AT %QB6544 : Byte;
   "SDC_EMS01_Carrier34_Zone" AT %QB6545 : Byte;
   "SDC_EMS01_Carrier35_Zone" AT %QB6546 : Byte;
   "SDC_EMS01_Carrier36_Zone" AT %QB6547 : Byte;
   "SDC_EMS01_Carrier37_Zone" AT %QB6548 : Byte;
   "SDC_EMS01_Carrier38_Zone" AT %QB6549 : Byte;
   "SDC_EMS01_Carrier39_Zone" AT %QB6550 : Byte;
   "SDC_EMS01_Carrier40_Zone" AT %QB6551 : Byte;
   "SDC_EMS01_Carrier41_Zone" AT %QB6552 : Byte;
   "SDC_EMS01_Carrier42_Zone" AT %QB6553 : Byte;
   "SDC_EMS01_Carrier43_Zone" AT %QB6554 : Byte;
   "SDC_EMS01_Carrier44_Zone" AT %QB6555 : Byte;
   "SDC_EMS01_Carrier45_Zone" AT %QB6556 : Byte;
   "SDC_EMS01_Carrier46_Zone" AT %QB6557 : Byte;
   "SDC_EMS01_Carrier47_Zone" AT %QB6558 : Byte;
   "SDC_EMS01_Carrier48_Zone" AT %QB6559 : Byte;
   "SDC_EMS01_Carrier49_Zone" AT %QB6560 : Byte;
   "SDC_EMS01_Carrier50_Zone" AT %QB6561 : Byte;
   "SDC_EMS01_Carrier51_Zone" AT %QB6562 : Byte;
   "SDC_EMS01_Carrier52_Zone" AT %QB6563 : Byte;
   "SDC_EMS01_Carrier53_Zone" AT %QB6564 : Byte;
   "SDC_EMS01_Carrier54_Zone" AT %QB6565 : Byte;
   "SDC_EMS01_Carrier55_Zone" AT %QB6566 : Byte;
   "SDC_EMS01_Carrier56_Zone" AT %QB6567 : Byte;
   "SDC_EMS01_Carrier57_Zone" AT %QB6568 : Byte;
   "SDC_EMS01_Carrier58_Zone" AT %QB6569 : Byte;
   "SDC_EMS01_Carrier59_Zone" AT %QB6570 : Byte;
   "SDC_EMS01_Carrier60_Zone" AT %QB6571 : Byte;
   "SDC_EMS01_Carrier61_Zone" AT %QB6572 : Byte;
   "SDC_EMS01_Carrier62_Zone" AT %QB6573 : Byte;
   "SDC_EMS01_Carrier63_Zone" AT %QB6574 : Byte;
   "SDC_EMS01_Carrier64_Zone" AT %QB6575 : Byte;
   "SDC_EMS01_Carrier65_Zone" AT %QB6576 : Byte;
   "SDC_EMS01_Carrier66_Zone" AT %QB6577 : Byte;
   "SDC_EMS01_Carrier67_Zone" AT %QB6578 : Byte;
   "SDC_EMS01_Carrier68_Zone" AT %QB6579 : Byte;
   "SDC_EMS01_Carrier69_Zone" AT %QB6580 : Byte;
   "SDC_EMS01_Carrier70_Zone" AT %QB6581 : Byte;
   "SDC_EMS01_Carrier71_Zone" AT %QB6582 : Byte;
   "SDC_EMS01_Carrier72_Zone" AT %QB6583 : Byte;
   "SDC_EMS01_Carrier73_Zone" AT %QB6584 : Byte;
   "SDC_EMS01_Carrier74_Zone" AT %QB6585 : Byte;
   "SDC_EMS01_Carrier75_Zone" AT %QB6586 : Byte;
   "SDC_EMS01_Carrier76_Zone" AT %QB6587 : Byte;
   "SDC_EMS01_Carrier77_Zone" AT %QB6588 : Byte;
   "SDC_EMS01_Carrier78_Zone" AT %QB6589 : Byte;
   "SDC_EMS01_Carrier79_Zone" AT %QB6590 : Byte;
   "SDC_EMS01_Carrier80_Zone" AT %QB6591 : Byte;
   "SDC_EMS01_Carrier81_Zone" AT %QB6592 : Byte;
   "SDC_EMS01_Carrier82_Zone" AT %QB6593 : Byte;
   "SDC_EMS01_Carrier83_Zone" AT %QB6594 : Byte;
   "SDC_EMS01_Carrier84_Zone" AT %QB6595 : Byte;
   "SDC_EMS01_Carrier85_Zone" AT %QB6596 : Byte;
   "SDC_EMS01_Carrier86_Zone" AT %QB6597 : Byte;
   "SDC_EMS01_Carrier87_Zone" AT %QB6598 : Byte;
   "SDC_EMS01_Carrier88_Zone" AT %QB6599 : Byte;
   "SDC_EMS01_Carrier89_Zone" AT %QB6600 : Byte;
   "SDC_EMS01_Carrier90_Zone" AT %QB6601 : Byte;
   "SDC_EMS01_Carrier91_Zone" AT %QB6602 : Byte;
   "SDC_EMS01_Carrier92_Zone" AT %QB6603 : Byte;
   "SDC_EMS01_Carrier93_Zone" AT %QB6604 : Byte;
   "SDC_EMS01_Carrier94_Zone" AT %QB6605 : Byte;
   "SDC_EMS01_Carrier95_Zone" AT %QB6606 : Byte;
   "SDC_EMS01_Carrier1_Position" AT %QD6000 : DWord;
   "SDC_EMS01_Carrier2_Position" AT %QD6004 : DWord;
   "SDC_EMS01_Carrier3_Position" AT %QD6008 : DWord;
   "SDC_EMS01_Carrier4_Position" AT %QD6012 : DWord;
   "SDC_EMS01_Carrier5_Position" AT %QD6016 : DWord;
   "SDC_EMS01_Carrier6_Position" AT %QD6020 : DWord;
   "SDC_EMS01_Carrier7_Position" AT %QD6024 : DWord;
   "SDC_EMS01_Carrier8_Position" AT %QD6028 : DWord;
   "SDC_EMS01_Carrier9_Position" AT %QD6032 : DWord;
   "SDC_EMS01_Carrier10_Position" AT %QD6036 : DWord;
   "SDC_EMS01_Carrier11_Position" AT %QD6040 : DWord;
   "SDC_EMS01_Carrier12_Position" AT %QD6044 : DWord;
   "SDC_EMS01_Carrier13_Position" AT %QD6048 : DWord;
   "SDC_EMS01_Carrier14_Position" AT %QD6052 : DWord;
   "SDC_EMS01_Carrier15_Position" AT %QD6056 : DWord;
   "SDC_EMS01_Carrier16_Position" AT %QD6060 : DWord;
   "SDC_EMS01_Carrier17_Position" AT %QD6064 : DWord;
   "SDC_EMS01_Carrier18_Position" AT %QD6068 : DWord;
   "SDC_EMS01_Carrier19_Position" AT %QD6072 : DWord;
   "SDC_EMS01_Carrier20_Position" AT %QD6076 : DWord;
   "SDC_EMS01_Carrier21_Position" AT %QD6080 : DWord;
   "SDC_EMS01_Carrier22_Position" AT %QD6084 : DWord;
   "SDC_EMS01_Carrier23_Position" AT %QD6088 : DWord;
   "SDC_EMS01_Carrier24_Position" AT %QD6092 : DWord;
   "SDC_EMS01_Carrier25_Position" AT %QD6096 : DWord;
   "SDC_EMS01_Carrier26_Position" AT %QD6100 : DWord;
   "SDC_EMS01_Carrier28_Position" AT %QD6108 : DWord;
   "SDC_EMS01_Carrier29_Position" AT %QD6112 : DWord;
   "SDC_EMS01_Carrier30_Position" AT %QD6116 : DWord;
   "SDC_EMS01_Carrier31_Position" AT %QD6120 : DWord;
   "SDC_EMS01_Carrier32_Position" AT %QD6124 : DWord;
   "SDC_EMS01_Carrier33_Position" AT %QD6128 : DWord;
   "SDC_EMS01_Carrier34_Position" AT %QD6132 : DWord;
   "SDC_EMS01_Carrier35_Position" AT %QD6136 : DWord;
   "SDC_EMS01_Carrier36_Position" AT %QD6140 : DWord;
   "SDC_EMS01_Carrier37_Position" AT %QD6144 : DWord;
   "SDC_EMS01_Carrier38_Position" AT %QD6148 : DWord;
   "SDC_EMS01_Carrier39_Position" AT %QD6152 : DWord;
   "SDC_EMS01_Carrier40_Position" AT %QD6156 : DWord;
   "SDC_EMS01_Carrier41_Position" AT %QD6160 : DWord;
   "SDC_EMS01_Carrier42_Position" AT %QD6164 : DWord;
   "SDC_EMS01_Carrier43_Position" AT %QD6168 : DWord;
   "SDC_EMS01_Carrier44_Position" AT %QD6172 : DWord;
   "SDC_EMS01_Carrier45_Position" AT %QD6176 : DWord;
   "SDC_EMS01_Carrier46_Position" AT %QD6180 : DWord;
   "SDC_EMS01_Carrier47_Position" AT %QD6184 : DWord;
   "SDC_EMS01_Carrier48_Position" AT %QD6188 : DWord;
   "SDC_EMS01_Carrier49_Position" AT %QD6192 : DWord;
   "SDC_EMS01_Carrier50_Position" AT %QD6196 : DWord;
   "SDC_EMS01_Carrier51_Position" AT %QD6200 : DWord;
   "SDC_EMS01_Carrier52_Position" AT %QD6204 : DWord;
   "SDC_EMS01_Carrier53_Position" AT %QD6208 : DWord;
   "SDC_EMS01_Carrier54_Position" AT %QD6212 : DWord;
   "SDC_EMS01_Carrier55_Position" AT %QD6216 : DWord;
   "SDC_EMS01_Carrier56_Position" AT %QD6220 : DWord;
   "SDC_EMS01_Carrier57_Position" AT %QD6224 : DWord;
   "SDC_EMS01_Carrier58_Position" AT %QD6228 : DWord;
   "SDC_EMS01_Carrier59_Position" AT %QD6232 : DWord;
   "SDC_EMS01_Carrier60_Position" AT %QD6236 : DWord;
   "SDC_EMS01_Carrier61_Position" AT %QD6240 : DWord;
   "SDC_EMS01_Carrier62_Position" AT %QD6244 : DWord;
   "SDC_EMS01_Carrier63_Position" AT %QD6248 : DWord;
   "SDC_EMS01_Carrier64_Position" AT %QD6252 : DWord;
   "SDC_EMS01_Carrier65_Position" AT %QD6256 : DWord;
   "SDC_EMS01_Carrier66_Position" AT %QD6260 : DWord;
   "SDC_EMS01_Carrier67_Position" AT %QD6264 : DWord;
   "SDC_EMS01_Carrier68_Position" AT %QD6268 : DWord;
   "SDC_EMS01_Carrier69_Position" AT %QD6272 : DWord;
   "SDC_EMS01_Carrier70_Position" AT %QD6276 : DWord;
   "SDC_EMS01_Carrier71_Position" AT %QD6280 : DWord;
   "SDC_EMS01_Carrier72_Position" AT %QD6284 : DWord;
   "SDC_EMS01_Carrier73_Position" AT %QD6288 : DWord;
   "SDC_EMS01_Carrier74_Position" AT %QD6292 : DWord;
   "SDC_EMS01_Carrier75_Position" AT %QD6296 : DWord;
   "SDC_EMS01_Carrier76_Position" AT %QD6300 : DWord;
   "SDC_EMS01_Carrier77_Position" AT %QD6304 : DWord;
   "SDC_EMS01_Carrier78_Position" AT %QD6308 : DWord;
   "SDC_EMS01_Carrier79_Position" AT %QD6312 : DWord;
   "SDC_EMS01_Carrier80_Position" AT %QD6316 : DWord;
   "SDC_EMS01_Carrier81_Position" AT %QD6320 : DWord;
   "SDC_EMS01_Carrier82_Position" AT %QD6324 : DWord;
   "SDC_EMS01_Carrier83_Position" AT %QD6328 : DWord;
   "SDC_EMS01_Carrier84_Position" AT %QD6332 : DWord;
   "SDC_EMS01_Carrier85_Position" AT %QD6336 : DWord;
   "SDC_EMS01_Carrier86_Position" AT %QD6340 : DWord;
   "SDC_EMS01_Carrier87_Position" AT %QD6344 : DWord;
   "SDC_EMS01_Carrier88_Position" AT %QD6348 : DWord;
   "SDC_EMS01_Carrier89_Position" AT %QD6352 : DWord;
   "SDC_EMS01_Carrier90_Position" AT %QD6356 : DWord;
   "SDC_EMS01_Carrier91_Position" AT %QD6360 : DWord;
   "SDC_EMS01_Carrier92_Position" AT %QD6364 : DWord;
   "SDC_EMS01_Carrier93_Position" AT %QD6368 : DWord;
   "SDC_EMS01_Carrier94_Position" AT %QD6372 : DWord;
   "SDC_EMS01_Carrier95_Position" AT %QD6376 : DWord;
END_VAR

